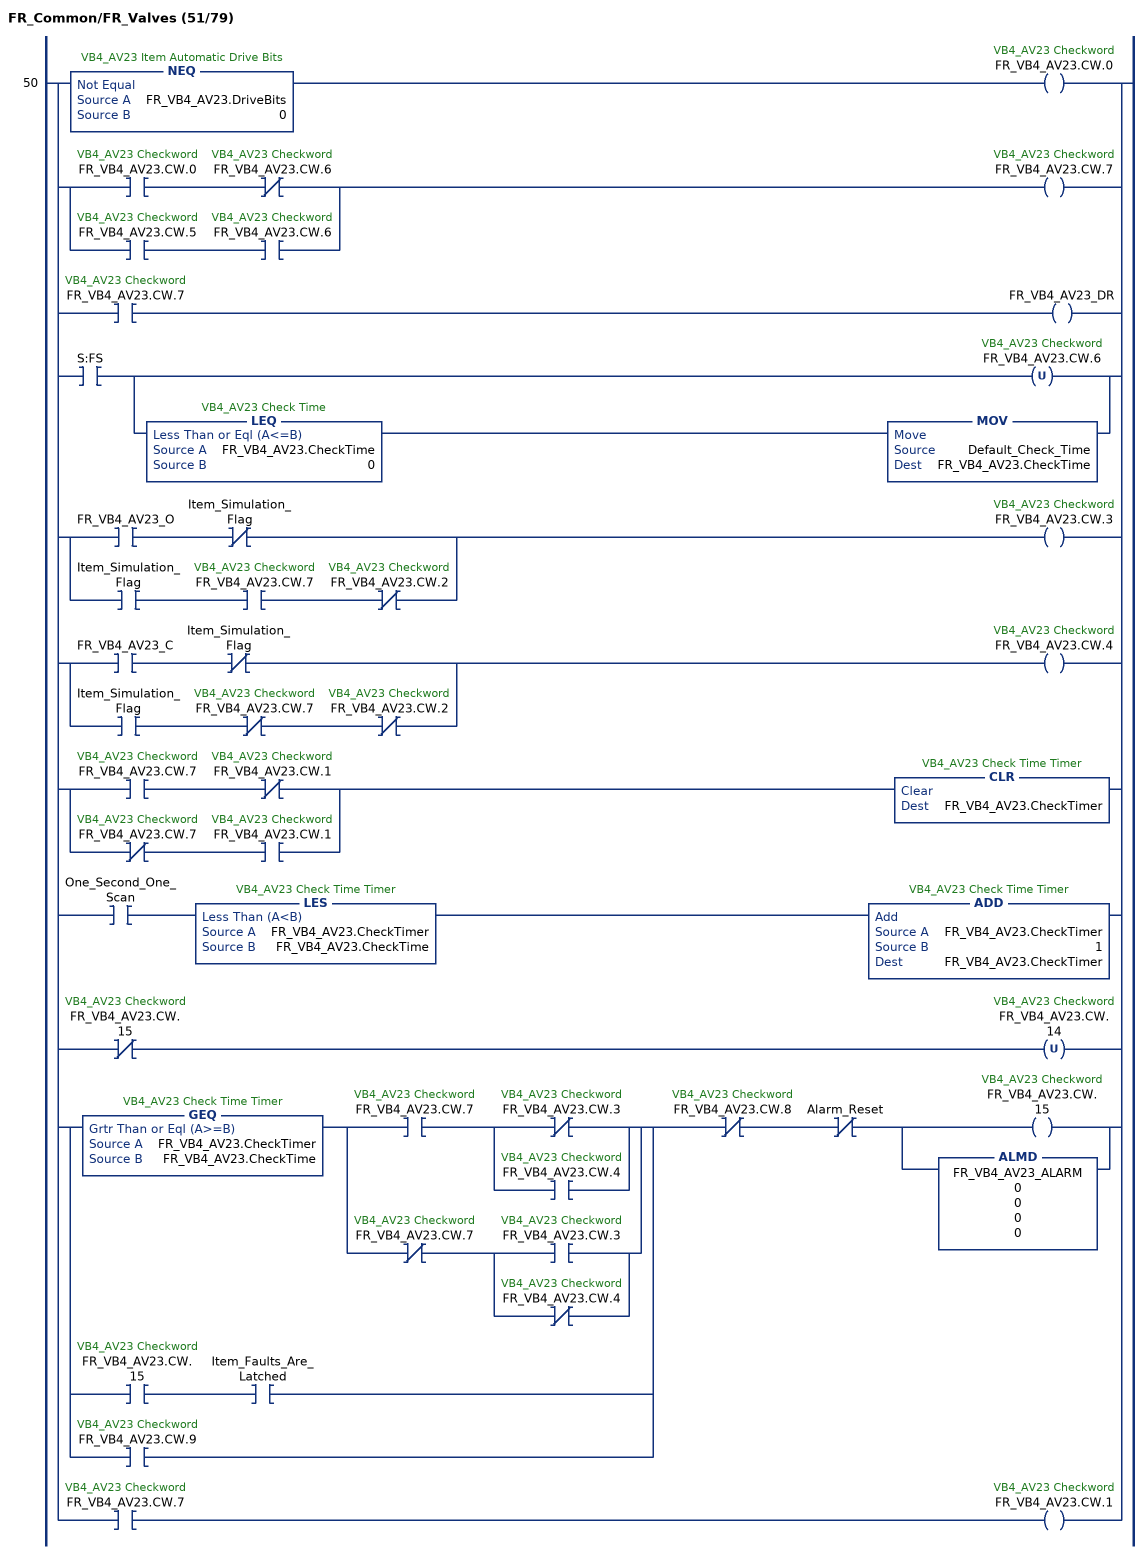
   50: [NEQ(FR_VB4_AV23.DriveBits,0) OTE(FR_VB4_AV23.CW.0) ,[XIC(FR_VB4_AV23.CW.0) XIO(FR_VB4_AV23.CW.6) ,XIC(FR_VB4_AV23.CW.5) XIC(FR_VB4_AV23.CW.6) ] OTE(FR_VB4_AV23.CW.7) ,XIC(FR_VB4_AV23.CW.7) OTE(FR_VB4_AV23_DR) ,XIC(S:FS) [OTU(FR_VB4_AV23.CW.6) ,LEQ(FR_VB4_AV23.CheckTime,0) MOV(Default_Check_Time,FR_VB4_AV23.CheckTime) ] ,[[XIC(FR_VB4_AV23_O) XIO(Item_Simulation_Flag) ,XIC(Item_Simulation_Flag) XIC(FR_VB4_AV23.CW.7) XIO(FR_VB4_AV23.CW.2) ] OTE(FR_VB4_AV23.CW.3) ,[XIC(FR_VB4_AV23_C) XIO(Item_Simulation_Flag) ,XIC(Item_Simulation_Flag) XIO(FR_VB4_AV23.CW.7) XIO(FR_VB4_AV23.CW.2) ] OTE(FR_VB4_AV23.CW.4) ] ,[XIC(FR_VB4_AV23.CW.7) XIO(FR_VB4_AV23.CW.1) ,XIO(FR_VB4_AV23.CW.7) XIC(FR_VB4_AV23.CW.1) ] CLR(FR_VB4_AV23.CheckTimer) ,XIC(One_Second_One_Scan) LES(FR_VB4_AV23.CheckTimer,FR_VB4_AV23.CheckTime) ADD(FR_VB4_AV23.CheckTimer,1,FR_VB4_AV23.CheckTimer) ,XIO(FR_VB4_AV23.CW.15) OTU(FR_VB4_AV23.CW.14) ,[GEQ(FR_VB4_AV23.CheckTimer,FR_VB4_AV23.CheckTime) [XIC(FR_VB4_AV23.CW.7) [XIO(FR_VB4_AV23.CW.3) ,XIC(FR_VB4_AV23.CW.4) ] ,XIO(FR_VB4_AV23.CW.7) [XIC(FR_VB4_AV23.CW.3) ,XIO(FR_VB4_AV23.CW.4) ] ] ,XIC(FR_VB4_AV23.CW.15) XIC(Item_Faults_Are_Latched) ,XIC(FR_VB4_AV23.CW.9) ] XIO(FR_VB4_AV23.CW.8) XIO(Alarm_Reset) [OTE(FR_VB4_AV23.CW.15) ,ALMD(FR_VB4_AV23_ALARM,0,0,0,0) ] ,XIC(FR_VB4_AV23.CW.7) OTE(FR_VB4_AV23.CW.1) ];
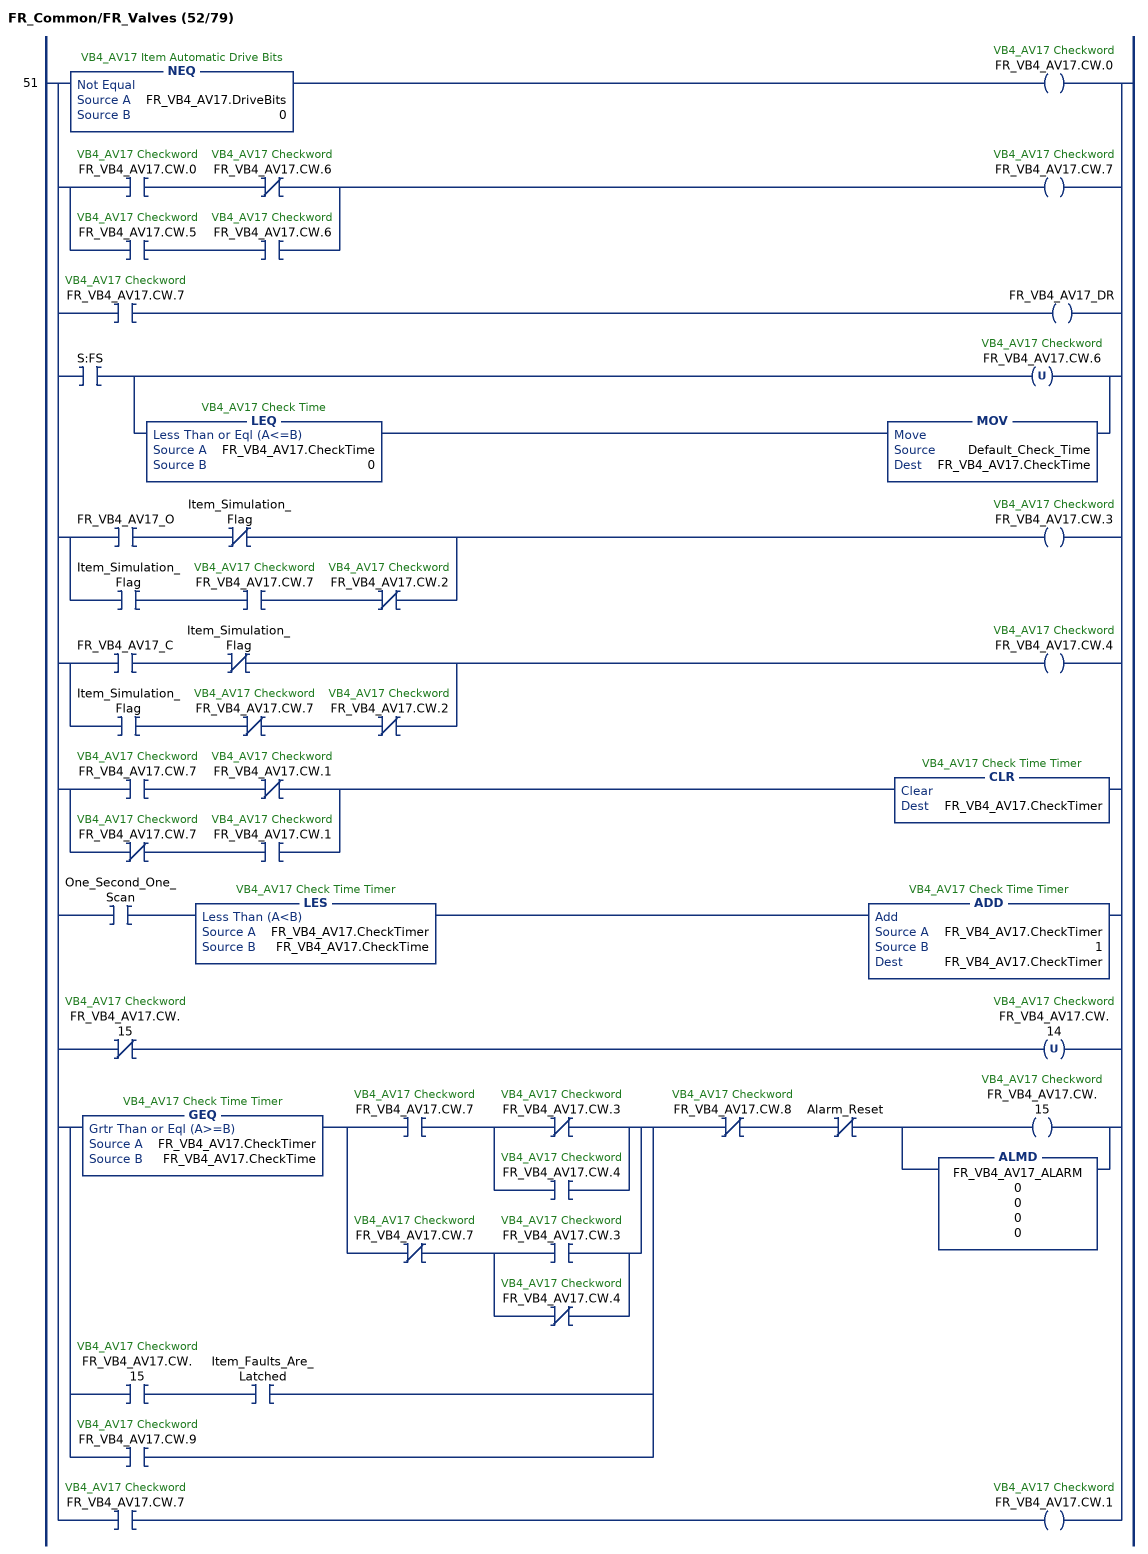
   51: [NEQ(FR_VB4_AV17.DriveBits,0) OTE(FR_VB4_AV17.CW.0) ,[XIC(FR_VB4_AV17.CW.0) XIO(FR_VB4_AV17.CW.6) ,XIC(FR_VB4_AV17.CW.5) XIC(FR_VB4_AV17.CW.6) ] OTE(FR_VB4_AV17.CW.7) ,XIC(FR_VB4_AV17.CW.7) OTE(FR_VB4_AV17_DR) ,XIC(S:FS) [OTU(FR_VB4_AV17.CW.6) ,LEQ(FR_VB4_AV17.CheckTime,0) MOV(Default_Check_Time,FR_VB4_AV17.CheckTime) ] ,[[XIC(FR_VB4_AV17_O) XIO(Item_Simulation_Flag) ,XIC(Item_Simulation_Flag) XIC(FR_VB4_AV17.CW.7) XIO(FR_VB4_AV17.CW.2) ] OTE(FR_VB4_AV17.CW.3) ,[XIC(FR_VB4_AV17_C) XIO(Item_Simulation_Flag) ,XIC(Item_Simulation_Flag) XIO(FR_VB4_AV17.CW.7) XIO(FR_VB4_AV17.CW.2) ] OTE(FR_VB4_AV17.CW.4) ] ,[XIC(FR_VB4_AV17.CW.7) XIO(FR_VB4_AV17.CW.1) ,XIO(FR_VB4_AV17.CW.7) XIC(FR_VB4_AV17.CW.1) ] CLR(FR_VB4_AV17.CheckTimer) ,XIC(One_Second_One_Scan) LES(FR_VB4_AV17.CheckTimer,FR_VB4_AV17.CheckTime) ADD(FR_VB4_AV17.CheckTimer,1,FR_VB4_AV17.CheckTimer) ,XIO(FR_VB4_AV17.CW.15) OTU(FR_VB4_AV17.CW.14) ,[GEQ(FR_VB4_AV17.CheckTimer,FR_VB4_AV17.CheckTime) [XIC(FR_VB4_AV17.CW.7) [XIO(FR_VB4_AV17.CW.3) ,XIC(FR_VB4_AV17.CW.4) ] ,XIO(FR_VB4_AV17.CW.7) [XIC(FR_VB4_AV17.CW.3) ,XIO(FR_VB4_AV17.CW.4) ] ] ,XIC(FR_VB4_AV17.CW.15) XIC(Item_Faults_Are_Latched) ,XIC(FR_VB4_AV17.CW.9) ] XIO(FR_VB4_AV17.CW.8) XIO(Alarm_Reset) [OTE(FR_VB4_AV17.CW.15) ,ALMD(FR_VB4_AV17_ALARM,0,0,0,0) ] ,XIC(FR_VB4_AV17.CW.7) OTE(FR_VB4_AV17.CW.1) ];
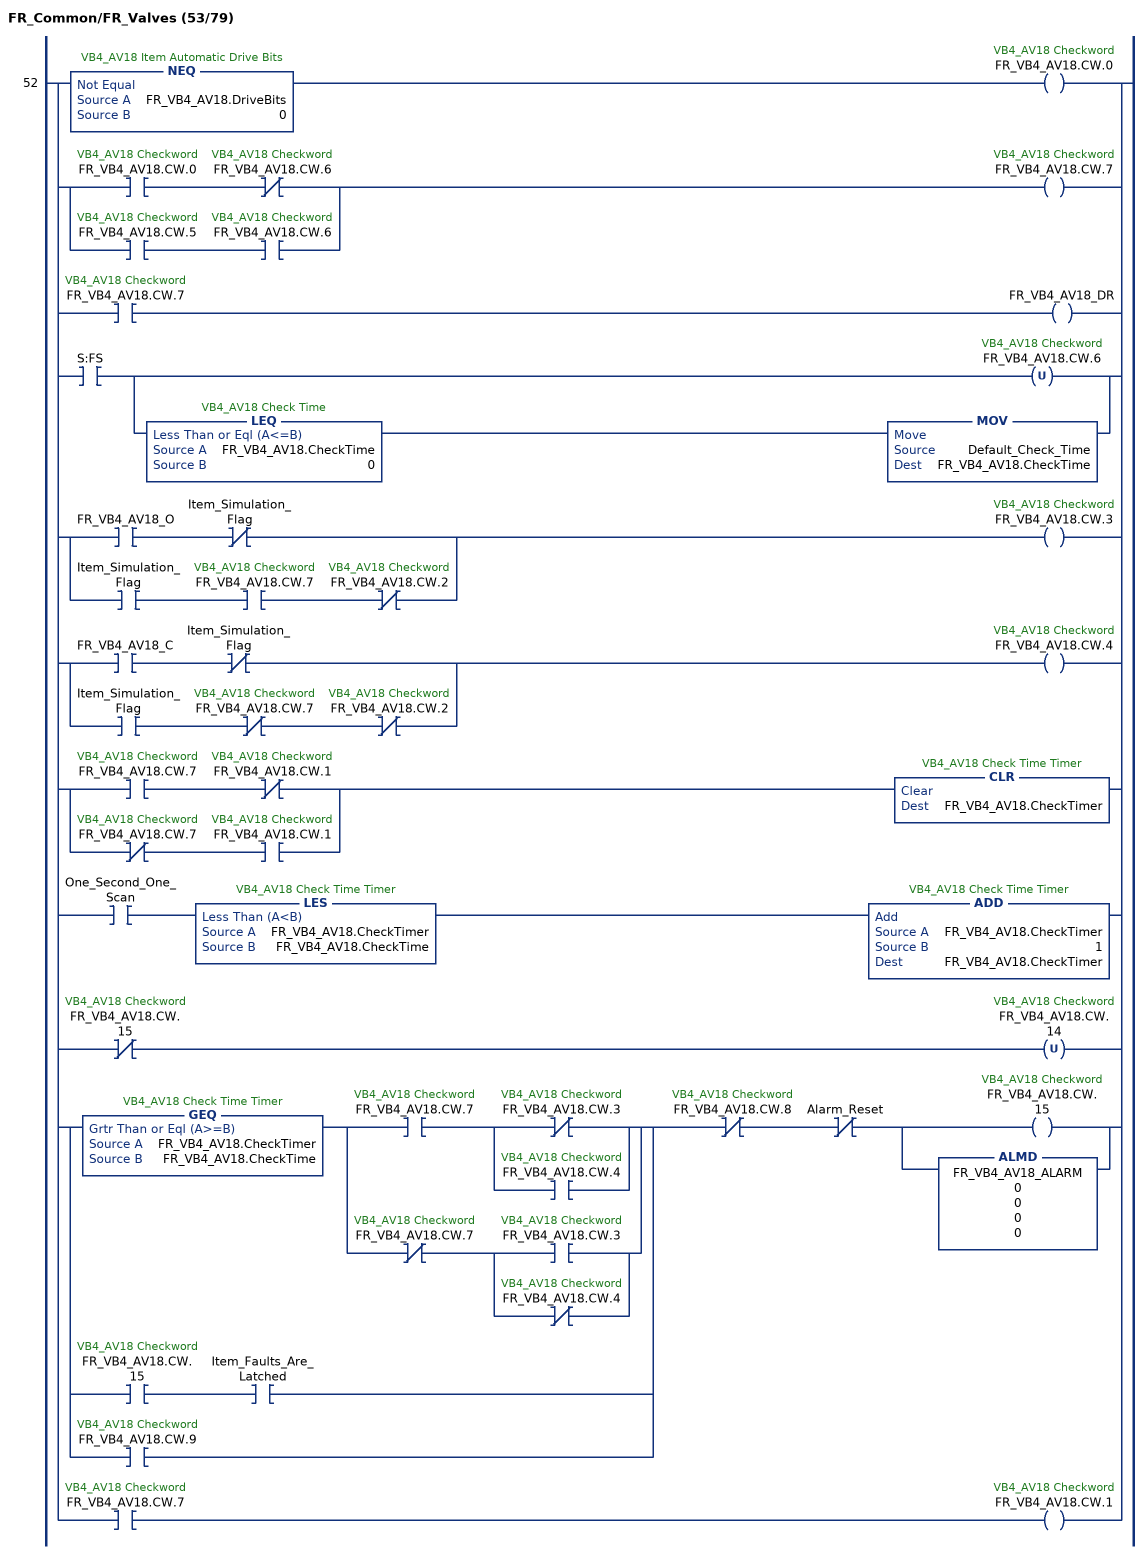
   52: [NEQ(FR_VB4_AV18.DriveBits,0) OTE(FR_VB4_AV18.CW.0) ,[XIC(FR_VB4_AV18.CW.0) XIO(FR_VB4_AV18.CW.6) ,XIC(FR_VB4_AV18.CW.5) XIC(FR_VB4_AV18.CW.6) ] OTE(FR_VB4_AV18.CW.7) ,XIC(FR_VB4_AV18.CW.7) OTE(FR_VB4_AV18_DR) ,XIC(S:FS) [OTU(FR_VB4_AV18.CW.6) ,LEQ(FR_VB4_AV18.CheckTime,0) MOV(Default_Check_Time,FR_VB4_AV18.CheckTime) ] ,[[XIC(FR_VB4_AV18_O) XIO(Item_Simulation_Flag) ,XIC(Item_Simulation_Flag) XIC(FR_VB4_AV18.CW.7) XIO(FR_VB4_AV18.CW.2) ] OTE(FR_VB4_AV18.CW.3) ,[XIC(FR_VB4_AV18_C) XIO(Item_Simulation_Flag) ,XIC(Item_Simulation_Flag) XIO(FR_VB4_AV18.CW.7) XIO(FR_VB4_AV18.CW.2) ] OTE(FR_VB4_AV18.CW.4) ] ,[XIC(FR_VB4_AV18.CW.7) XIO(FR_VB4_AV18.CW.1) ,XIO(FR_VB4_AV18.CW.7) XIC(FR_VB4_AV18.CW.1) ] CLR(FR_VB4_AV18.CheckTimer) ,XIC(One_Second_One_Scan) LES(FR_VB4_AV18.CheckTimer,FR_VB4_AV18.CheckTime) ADD(FR_VB4_AV18.CheckTimer,1,FR_VB4_AV18.CheckTimer) ,XIO(FR_VB4_AV18.CW.15) OTU(FR_VB4_AV18.CW.14) ,[GEQ(FR_VB4_AV18.CheckTimer,FR_VB4_AV18.CheckTime) [XIC(FR_VB4_AV18.CW.7) [XIO(FR_VB4_AV18.CW.3) ,XIC(FR_VB4_AV18.CW.4) ] ,XIO(FR_VB4_AV18.CW.7) [XIC(FR_VB4_AV18.CW.3) ,XIO(FR_VB4_AV18.CW.4) ] ] ,XIC(FR_VB4_AV18.CW.15) XIC(Item_Faults_Are_Latched) ,XIC(FR_VB4_AV18.CW.9) ] XIO(FR_VB4_AV18.CW.8) XIO(Alarm_Reset) [OTE(FR_VB4_AV18.CW.15) ,ALMD(FR_VB4_AV18_ALARM,0,0,0,0) ] ,XIC(FR_VB4_AV18.CW.7) OTE(FR_VB4_AV18.CW.1) ];
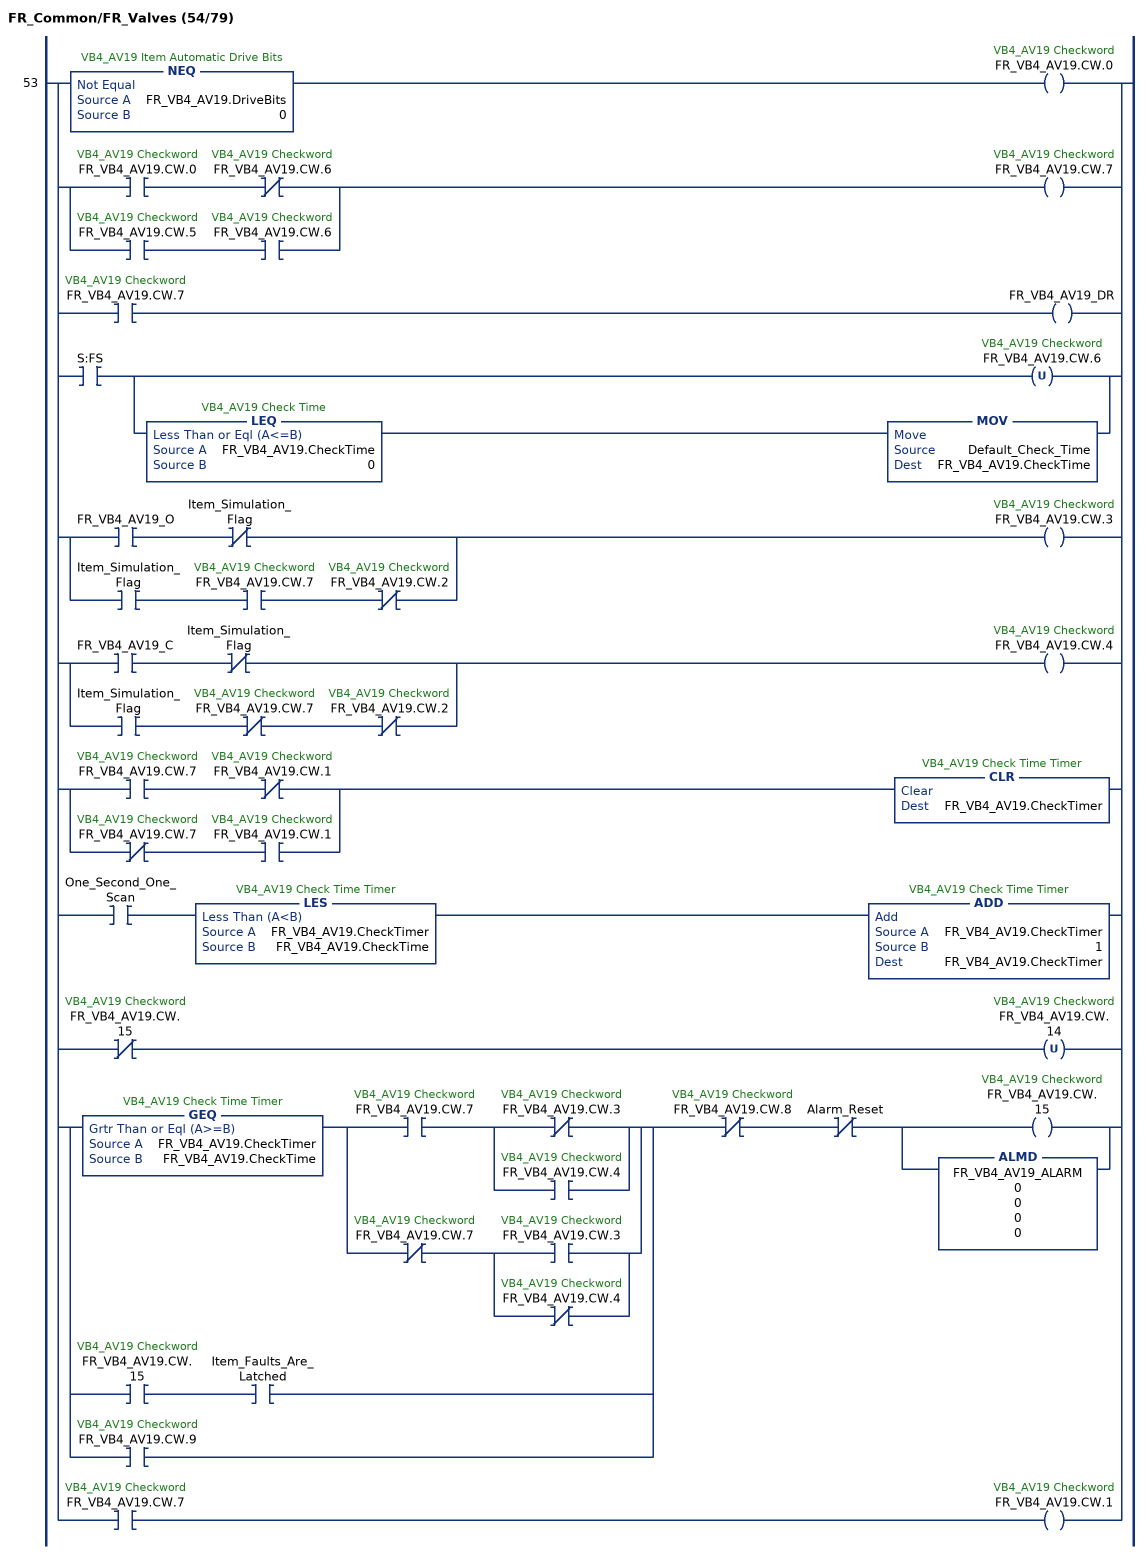
   53: [NEQ(FR_VB4_AV19.DriveBits,0) OTE(FR_VB4_AV19.CW.0) ,[XIC(FR_VB4_AV19.CW.0) XIO(FR_VB4_AV19.CW.6) ,XIC(FR_VB4_AV19.CW.5) XIC(FR_VB4_AV19.CW.6) ] OTE(FR_VB4_AV19.CW.7) ,XIC(FR_VB4_AV19.CW.7) OTE(FR_VB4_AV19_DR) ,XIC(S:FS) [OTU(FR_VB4_AV19.CW.6) ,LEQ(FR_VB4_AV19.CheckTime,0) MOV(Default_Check_Time,FR_VB4_AV19.CheckTime) ] ,[[XIC(FR_VB4_AV19_O) XIO(Item_Simulation_Flag) ,XIC(Item_Simulation_Flag) XIC(FR_VB4_AV19.CW.7) XIO(FR_VB4_AV19.CW.2) ] OTE(FR_VB4_AV19.CW.3) ,[XIC(FR_VB4_AV19_C) XIO(Item_Simulation_Flag) ,XIC(Item_Simulation_Flag) XIO(FR_VB4_AV19.CW.7) XIO(FR_VB4_AV19.CW.2) ] OTE(FR_VB4_AV19.CW.4) ] ,[XIC(FR_VB4_AV19.CW.7) XIO(FR_VB4_AV19.CW.1) ,XIO(FR_VB4_AV19.CW.7) XIC(FR_VB4_AV19.CW.1) ] CLR(FR_VB4_AV19.CheckTimer) ,XIC(One_Second_One_Scan) LES(FR_VB4_AV19.CheckTimer,FR_VB4_AV19.CheckTime) ADD(FR_VB4_AV19.CheckTimer,1,FR_VB4_AV19.CheckTimer) ,XIO(FR_VB4_AV19.CW.15) OTU(FR_VB4_AV19.CW.14) ,[GEQ(FR_VB4_AV19.CheckTimer,FR_VB4_AV19.CheckTime) [XIC(FR_VB4_AV19.CW.7) [XIO(FR_VB4_AV19.CW.3) ,XIC(FR_VB4_AV19.CW.4) ] ,XIO(FR_VB4_AV19.CW.7) [XIC(FR_VB4_AV19.CW.3) ,XIO(FR_VB4_AV19.CW.4) ] ] ,XIC(FR_VB4_AV19.CW.15) XIC(Item_Faults_Are_Latched) ,XIC(FR_VB4_AV19.CW.9) ] XIO(FR_VB4_AV19.CW.8) XIO(Alarm_Reset) [OTE(FR_VB4_AV19.CW.15) ,ALMD(FR_VB4_AV19_ALARM,0,0,0,0) ] ,XIC(FR_VB4_AV19.CW.7) OTE(FR_VB4_AV19.CW.1) ];
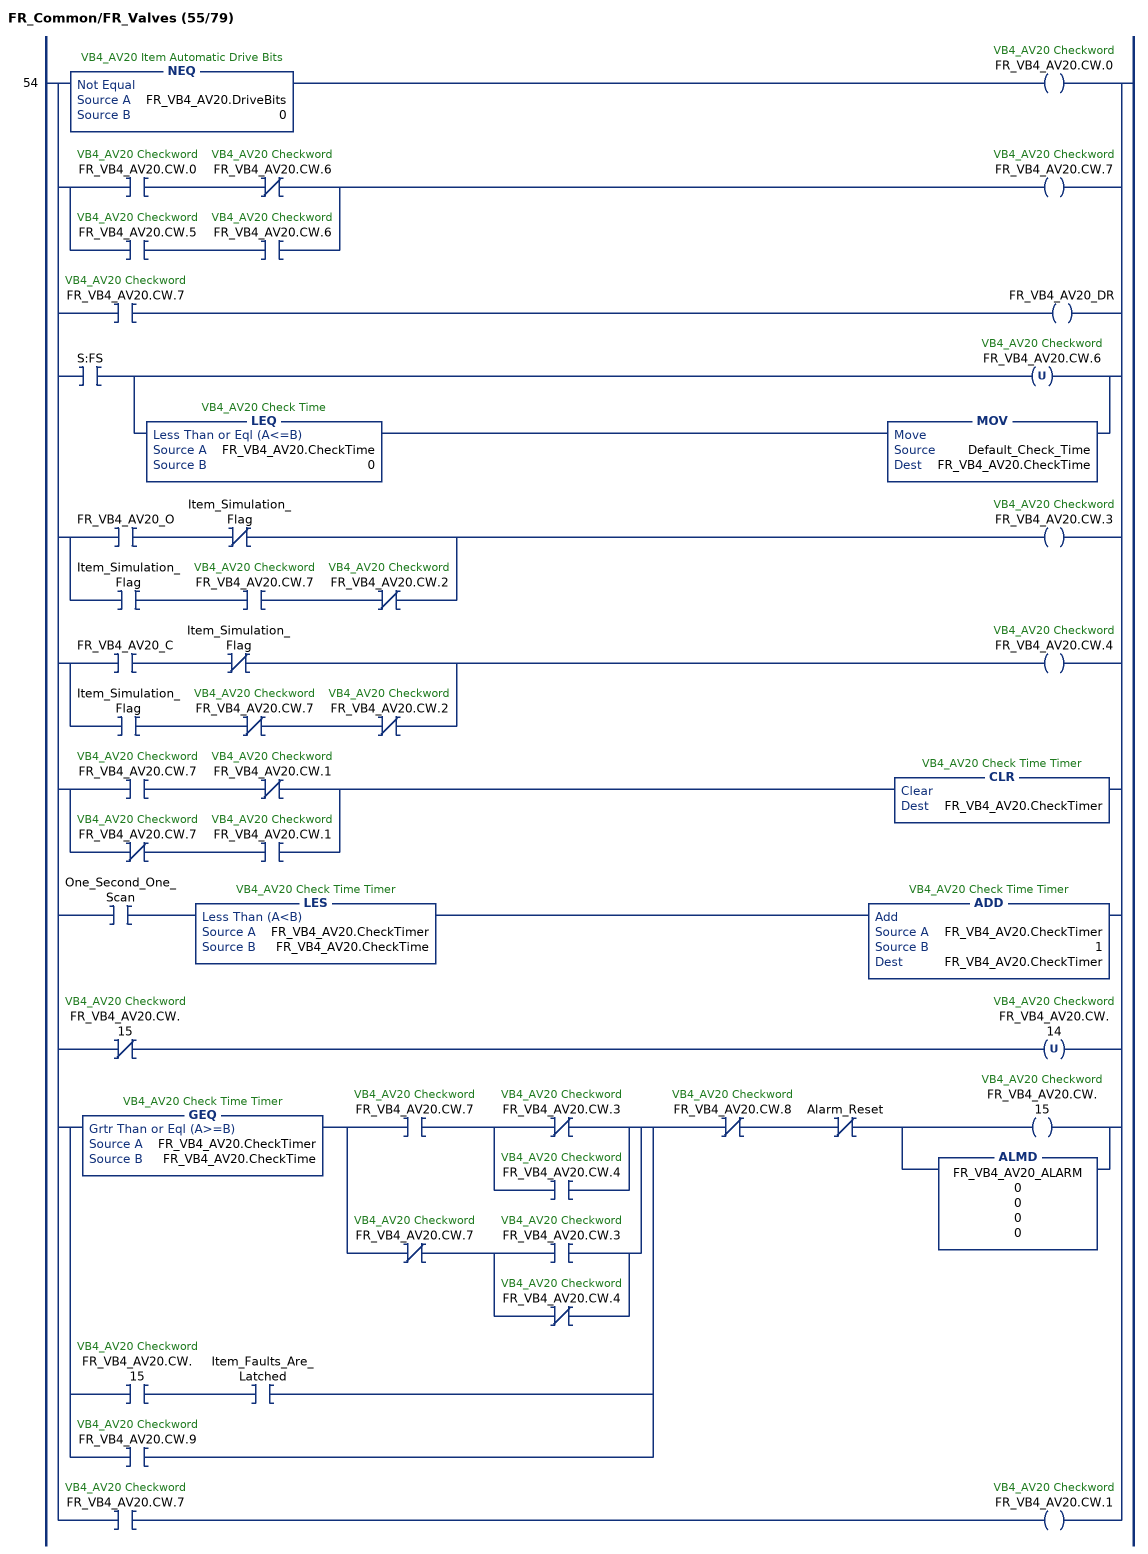
   54: [NEQ(FR_VB4_AV20.DriveBits,0) OTE(FR_VB4_AV20.CW.0) ,[XIC(FR_VB4_AV20.CW.0) XIO(FR_VB4_AV20.CW.6) ,XIC(FR_VB4_AV20.CW.5) XIC(FR_VB4_AV20.CW.6) ] OTE(FR_VB4_AV20.CW.7) ,XIC(FR_VB4_AV20.CW.7) OTE(FR_VB4_AV20_DR) ,XIC(S:FS) [OTU(FR_VB4_AV20.CW.6) ,LEQ(FR_VB4_AV20.CheckTime,0) MOV(Default_Check_Time,FR_VB4_AV20.CheckTime) ] ,[[XIC(FR_VB4_AV20_O) XIO(Item_Simulation_Flag) ,XIC(Item_Simulation_Flag) XIC(FR_VB4_AV20.CW.7) XIO(FR_VB4_AV20.CW.2) ] OTE(FR_VB4_AV20.CW.3) ,[XIC(FR_VB4_AV20_C) XIO(Item_Simulation_Flag) ,XIC(Item_Simulation_Flag) XIO(FR_VB4_AV20.CW.7) XIO(FR_VB4_AV20.CW.2) ] OTE(FR_VB4_AV20.CW.4) ] ,[XIC(FR_VB4_AV20.CW.7) XIO(FR_VB4_AV20.CW.1) ,XIO(FR_VB4_AV20.CW.7) XIC(FR_VB4_AV20.CW.1) ] CLR(FR_VB4_AV20.CheckTimer) ,XIC(One_Second_One_Scan) LES(FR_VB4_AV20.CheckTimer,FR_VB4_AV20.CheckTime) ADD(FR_VB4_AV20.CheckTimer,1,FR_VB4_AV20.CheckTimer) ,XIO(FR_VB4_AV20.CW.15) OTU(FR_VB4_AV20.CW.14) ,[GEQ(FR_VB4_AV20.CheckTimer,FR_VB4_AV20.CheckTime) [XIC(FR_VB4_AV20.CW.7) [XIO(FR_VB4_AV20.CW.3) ,XIC(FR_VB4_AV20.CW.4) ] ,XIO(FR_VB4_AV20.CW.7) [XIC(FR_VB4_AV20.CW.3) ,XIO(FR_VB4_AV20.CW.4) ] ] ,XIC(FR_VB4_AV20.CW.15) XIC(Item_Faults_Are_Latched) ,XIC(FR_VB4_AV20.CW.9) ] XIO(FR_VB4_AV20.CW.8) XIO(Alarm_Reset) [OTE(FR_VB4_AV20.CW.15) ,ALMD(FR_VB4_AV20_ALARM,0,0,0,0) ] ,XIC(FR_VB4_AV20.CW.7) OTE(FR_VB4_AV20.CW.1) ];